HMI tags "Tool_Editor"
   "DB_MouldEditor_HMI_uData_sSelected_iCalculation" : Int = PLC DB_MouldEditor_HMI.uData.sSelected.iCalculation AT %DB10.DBW92, 1 s
   "DB_MouldEditor_HMI_uData_arShotSet{1}_CPMoveAfterShot" : Bool = PLC DB_MouldEditor_HMI.uData.arShotSet[1].CPMoveAfterShot AT %DB10.DBX236.1, 1 s
   "DB_MouldEditor_HMI_uData_arShotSet{2}_CPMoveAfterShot" : Bool = PLC DB_MouldEditor_HMI.uData.arShotSet[2].CPMoveAfterShot AT %DB10.DBX308.1, 1 s
   "DB_MouldEditor_HMI_uData_arShotSet{3}_CPMoveAfterShot" : Bool = PLC DB_MouldEditor_HMI.uData.arShotSet[3].CPMoveAfterShot AT %DB10.DBX380.1, 1 s
   "DB_MouldEditor_HMI_uData_arShotSet{4}_CPMoveAfterShot" : Bool = PLC DB_MouldEditor_HMI.uData.arShotSet[4].CPMoveAfterShot AT %DB10.DBX452.1, 1 s
   "DB_MouldEditor_HMI_uData_arShotSet{5}_CPMoveAfterShot" : Bool = PLC DB_MouldEditor_HMI.uData.arShotSet[5].CPMoveAfterShot AT %DB10.DBX524.1, 1 s
   "DB_MouldEditor_HMI_uData_arShotSet{6}_CPMoveAfterShot" : Bool = PLC DB_MouldEditor_HMI.uData.arShotSet[6].CPMoveAfterShot AT %DB10.DBX596.1, 1 s
   "DB_MouldEditor_HMI_uData_arShotSet{7}_CPMoveAfterShot" : Bool = PLC DB_MouldEditor_HMI.uData.arShotSet[7].CPMoveAfterShot AT %DB10.DBX668.1, 1 s
   "DB_MouldEditor_HMI_uData_arShotSet{8}_CPMoveAfterShot" : Bool = PLC DB_MouldEditor_HMI.uData.arShotSet[8].CPMoveAfterShot AT %DB10.DBX740.1, 1 s
   "DB_MouldEditor_HMI_uData_uTools_EnableTool" : Bool = PLC DB_MouldEditor_HMI.uData.uTools.EnableTool AT %DB10.DBX771.0, 1 s
   "DB_MouldEditor_HMI_uData_sSelected_sPS_arFlow{1}" : Real = PLC DB_MouldEditor_HMI.uData.sSelected.sPS.arFlow[1] AT %DB10.DBD8, 1 s
   "DB_MouldEditor_HMI_uData_sSelected_sPS_arFlow{2}" : Real = PLC DB_MouldEditor_HMI.uData.sSelected.sPS.arFlow[2] AT %DB10.DBD12, 1 s
   "DB_MouldEditor_HMI_uData_sSelected_sPS_arFlow{3}" : Real = PLC DB_MouldEditor_HMI.uData.sSelected.sPS.arFlow[3] AT %DB10.DBD16, 1 s
   "DB_MouldEditor_HMI_uData_sSelected_sPS_arFlow{4}" : Real = PLC DB_MouldEditor_HMI.uData.sSelected.sPS.arFlow[4] AT %DB10.DBD20, 1 s
   "DB_MouldEditor_HMI_uData_sSelected_sPS_arFlow{5}" : Real = PLC DB_MouldEditor_HMI.uData.sSelected.sPS.arFlow[5] AT %DB10.DBD24, 1 s
   "DB_MouldEditor_HMI_uData_sSelected_sPS_arFlow{6}" : Real = PLC DB_MouldEditor_HMI.uData.sSelected.sPS.arFlow[6] AT %DB10.DBD28, 1 s
   "DB_MouldEditor_HMI_uData_arShotSet{1}_MHNo" : Int = PLC DB_MouldEditor_HMI.uData.arShotSet[1].MHNo AT %DB10.DBW166, 1 s
   "DB_MouldEditor_HMI_uData_arShotSet{2}_MHNo" : Int = PLC DB_MouldEditor_HMI.uData.arShotSet[2].MHNo AT %DB10.DBW238, 1 s
   "DB_MouldEditor_HMI_uData_arShotSet{3}_MHNo" : Int = PLC DB_MouldEditor_HMI.uData.arShotSet[3].MHNo AT %DB10.DBW310, 1 s
   "DB_MouldEditor_HMI_uData_arShotSet{4}_MHNo" : Int = PLC DB_MouldEditor_HMI.uData.arShotSet[4].MHNo AT %DB10.DBW382, 1 s
   "DB_MouldEditor_HMI_uData_arShotSet{5}_MHNo" : Int = PLC DB_MouldEditor_HMI.uData.arShotSet[5].MHNo AT %DB10.DBW454, 1 s
   "DB_MouldEditor_HMI_uData_arShotSet{6}_MHNo" : Int = PLC DB_MouldEditor_HMI.uData.arShotSet[6].MHNo AT %DB10.DBW526, 1 s
   "DB_MouldEditor_HMI_uData_arShotSet{7}_MHNo" : Int = PLC DB_MouldEditor_HMI.uData.arShotSet[7].MHNo AT %DB10.DBW598, 1 s
   "DB_MouldEditor_HMI_uData_arShotSet{8}_MHNo" : Int = PLC DB_MouldEditor_HMI.uData.arShotSet[8].MHNo AT %DB10.DBW670, 1 s
   "DB_MouldEditor_HMI_uData_arShotSet{1}_PartCounter" : Int = PLC DB_MouldEditor_HMI.uData.arShotSet[1].PartCounter AT %DB10.DBW184, 1 s
   "DB_MouldEditor_HMI_uData_arShotSet{2}_PartCounter" : Int = PLC DB_MouldEditor_HMI.uData.arShotSet[2].PartCounter AT %DB10.DBW256, 1 s
   "DB_MouldEditor_HMI_uData_arShotSet{3}_PartCounter" : Int = PLC DB_MouldEditor_HMI.uData.arShotSet[3].PartCounter AT %DB10.DBW328, 1 s
   "DB_MouldEditor_HMI_uData_arShotSet{4}_PartCounter" : Int = PLC DB_MouldEditor_HMI.uData.arShotSet[4].PartCounter AT %DB10.DBW400, 1 s
   "DB_MouldEditor_HMI_uData_arShotSet{5}_PartCounter" : Int = PLC DB_MouldEditor_HMI.uData.arShotSet[5].PartCounter AT %DB10.DBW472, 1 s
   "DB_MouldEditor_HMI_uData_arShotSet{6}_PartCounter" : Int = PLC DB_MouldEditor_HMI.uData.arShotSet[6].PartCounter AT %DB10.DBW544, 1 s
   "DB_MouldEditor_HMI_uData_arShotSet{7}_PartCounter" : Int = PLC DB_MouldEditor_HMI.uData.arShotSet[7].PartCounter AT %DB10.DBW616, 1 s
   "DB_MouldEditor_HMI_uData_arShotSet{8}_PartCounter" : Int = PLC DB_MouldEditor_HMI.uData.arShotSet[8].PartCounter AT %DB10.DBW688, 1 s
   "DB_MouldEditor_HMI_uData_arShotSet{1}_PartWeight" : Real = PLC DB_MouldEditor_HMI.uData.arShotSet[1].PartWeight AT %DB10.DBD172, 1 s
   "DB_MouldEditor_HMI_uData_arShotSet{2}_PartWeight" : Real = PLC DB_MouldEditor_HMI.uData.arShotSet[2].PartWeight AT %DB10.DBD244, 1 s
   "DB_MouldEditor_HMI_uData_arShotSet{3}_PartWeight" : Real = PLC DB_MouldEditor_HMI.uData.arShotSet[3].PartWeight AT %DB10.DBD316, 1 s
   "DB_MouldEditor_HMI_uData_arShotSet{4}_PartWeight" : Real = PLC DB_MouldEditor_HMI.uData.arShotSet[4].PartWeight AT %DB10.DBD388, 1 s
   "DB_MouldEditor_HMI_uData_arShotSet{5}_PartWeight" : Real = PLC DB_MouldEditor_HMI.uData.arShotSet[5].PartWeight AT %DB10.DBD460, 1 s
   "DB_MouldEditor_HMI_uData_arShotSet{6}_PartWeight" : Real = PLC DB_MouldEditor_HMI.uData.arShotSet[6].PartWeight AT %DB10.DBD532, 1 s
   "DB_MouldEditor_HMI_uData_arShotSet{7}_PartWeight" : Real = PLC DB_MouldEditor_HMI.uData.arShotSet[7].PartWeight AT %DB10.DBD604, 1 s
   "DB_MouldEditor_HMI_uData_arShotSet{8}_PartWeight" : Real = PLC DB_MouldEditor_HMI.uData.arShotSet[8].PartWeight AT %DB10.DBD676, 1 s
   "DB_MouldEditor_HMI_uData_sSelected_sPS_arPressure{1}" : Real = PLC DB_MouldEditor_HMI.uData.sSelected.sPS.arPressure[1] AT %DB10.DBD64, 1 s
   "DB_MouldEditor_HMI_uData_sSelected_sPS_arPressure{2}" : Real = PLC DB_MouldEditor_HMI.uData.sSelected.sPS.arPressure[2] AT %DB10.DBD68, 1 s
   "DB_MouldEditor_HMI_uData_sSelected_sPS_arPressure{3}" : Real = PLC DB_MouldEditor_HMI.uData.sSelected.sPS.arPressure[3] AT %DB10.DBD72, 1 s
   "DB_MouldEditor_HMI_uData_sSelected_sPS_arPressure{4}" : Real = PLC DB_MouldEditor_HMI.uData.sSelected.sPS.arPressure[4] AT %DB10.DBD76, 1 s
   "DB_MouldEditor_HMI_uData_sSelected_sPS_arPressure{5}" : Real = PLC DB_MouldEditor_HMI.uData.sSelected.sPS.arPressure[5] AT %DB10.DBD80, 1 s
   "DB_MouldEditor_HMI_uData_sSelected_sPS_arPressure{6}" : Real = PLC DB_MouldEditor_HMI.uData.sSelected.sPS.arPressure[6] AT %DB10.DBD84, 1 s
   "DB_MouldEditor_HMI_uData_arShotSet{1}_PartShotDisable" : Bool = PLC DB_MouldEditor_HMI.uData.arShotSet[1].PartShotDisable AT %DB10.DBX236.0, 1 s
   "DB_MouldEditor_HMI_uData_arShotSet{2}_PartShotDisable" : Bool = PLC DB_MouldEditor_HMI.uData.arShotSet[2].PartShotDisable AT %DB10.DBX308.0, 1 s
   "DB_MouldEditor_HMI_uData_arShotSet{3}_PartShotDisable" : Bool = PLC DB_MouldEditor_HMI.uData.arShotSet[3].PartShotDisable AT %DB10.DBX380.0, 1 s
   "DB_MouldEditor_HMI_uData_arShotSet{4}_PartShotDisable" : Bool = PLC DB_MouldEditor_HMI.uData.arShotSet[4].PartShotDisable AT %DB10.DBX452.0, 1 s
   "DB_MouldEditor_HMI_uData_arShotSet{5}_PartShotDisable" : Bool = PLC DB_MouldEditor_HMI.uData.arShotSet[5].PartShotDisable AT %DB10.DBX524.0, 1 s
   "DB_MouldEditor_HMI_uData_arShotSet{6}_PartShotDisable" : Bool = PLC DB_MouldEditor_HMI.uData.arShotSet[6].PartShotDisable AT %DB10.DBX596.0, 1 s
   "DB_MouldEditor_HMI_uData_arShotSet{7}_PartShotDisable" : Bool = PLC DB_MouldEditor_HMI.uData.arShotSet[7].PartShotDisable AT %DB10.DBX668.0, 1 s
   "DB_MouldEditor_HMI_uData_arShotSet{8}_PartShotDisable" : Bool = PLC DB_MouldEditor_HMI.uData.arShotSet[8].PartShotDisable AT %DB10.DBX740.0, 1 s
   "DB_MouldEditor_HMI_uData_sSelected_sPS_iPS" : Int = PLC DB_MouldEditor_HMI.uData.sSelected.sPS.iPS AT %DB10.DBW2, 1 s
   "DB_MouldEditor_HMI_uData_sSelected_sPS_arRatio{1}" : Real = PLC DB_MouldEditor_HMI.uData.sSelected.sPS.arRatio[1] AT %DB10.DBD36, 1 s
   "DB_MouldEditor_HMI_uData_sSelected_sPS_arRatio{2}" : Real = PLC DB_MouldEditor_HMI.uData.sSelected.sPS.arRatio[2] AT %DB10.DBD40, 1 s
   "DB_MouldEditor_HMI_uData_sSelected_sPS_arRatio{3}" : Real = PLC DB_MouldEditor_HMI.uData.sSelected.sPS.arRatio[3] AT %DB10.DBD44, 1 s
   "DB_MouldEditor_HMI_uData_sSelected_sPS_arRatio{4}" : Real = PLC DB_MouldEditor_HMI.uData.sSelected.sPS.arRatio[4] AT %DB10.DBD48, 1 s
   "DB_MouldEditor_HMI_uData_sSelected_sPS_arRatio{5}" : Real = PLC DB_MouldEditor_HMI.uData.sSelected.sPS.arRatio[5] AT %DB10.DBD52, 1 s
   "DB_MouldEditor_HMI_uData_sSelected_sPS_arRatio{6}" : Real = PLC DB_MouldEditor_HMI.uData.sSelected.sPS.arRatio[6] AT %DB10.DBD56, 1 s
   "DB_MouldEditor_HMI_uData_arShotSet{1}_PurgeMHAfterShot" : Bool = PLC DB_MouldEditor_HMI.uData.arShotSet[1].PurgeMHAfterShot AT %DB10.DBX236.2, 1 s
   "DB_MouldEditor_HMI_uData_arShotSet{2}_PurgeMHAfterShot" : Bool = PLC DB_MouldEditor_HMI.uData.arShotSet[2].PurgeMHAfterShot AT %DB10.DBX308.2, 1 s
   "DB_MouldEditor_HMI_uData_arShotSet{3}_PurgeMHAfterShot" : Bool = PLC DB_MouldEditor_HMI.uData.arShotSet[3].PurgeMHAfterShot AT %DB10.DBX380.2, 1 s
   "DB_MouldEditor_HMI_uData_arShotSet{4}_PurgeMHAfterShot" : Bool = PLC DB_MouldEditor_HMI.uData.arShotSet[4].PurgeMHAfterShot AT %DB10.DBX452.2, 1 s
   "DB_MouldEditor_HMI_uData_arShotSet{5}_PurgeMHAfterShot" : Bool = PLC DB_MouldEditor_HMI.uData.arShotSet[5].PurgeMHAfterShot AT %DB10.DBX524.2, 1 s
   "DB_MouldEditor_HMI_uData_arShotSet{6}_PurgeMHAfterShot" : Bool = PLC DB_MouldEditor_HMI.uData.arShotSet[6].PurgeMHAfterShot AT %DB10.DBX596.2, 1 s
   "DB_MouldEditor_HMI_uData_arShotSet{7}_PurgeMHAfterShot" : Bool = PLC DB_MouldEditor_HMI.uData.arShotSet[7].PurgeMHAfterShot AT %DB10.DBX668.2, 1 s
   "DB_MouldEditor_HMI_uData_arShotSet{8}_PurgeMHAfterShot" : Bool = PLC DB_MouldEditor_HMI.uData.arShotSet[8].PurgeMHAfterShot AT %DB10.DBX740.2, 1 s
   "DB_MouldEditor_HMI_uData_arShotSet{1}_FoamingTime" : Real = PLC DB_MouldEditor_HMI.uData.arShotSet[1].FoamingTime AT %DB10.DBD168, 1 s
   "DB_MouldEditor_HMI_uData_arShotSet{2}_FoamingTime" : Real = PLC DB_MouldEditor_HMI.uData.arShotSet[2].FoamingTime AT %DB10.DBD240, 1 s
   "DB_MouldEditor_HMI_uData_arShotSet{3}_FoamingTime" : Real = PLC DB_MouldEditor_HMI.uData.arShotSet[3].FoamingTime AT %DB10.DBD312, 1 s
   "DB_MouldEditor_HMI_uData_arShotSet{4}_FoamingTime" : Real = PLC DB_MouldEditor_HMI.uData.arShotSet[4].FoamingTime AT %DB10.DBD384, 1 s
   "DB_MouldEditor_HMI_uData_arShotSet{5}_FoamingTime" : Real = PLC DB_MouldEditor_HMI.uData.arShotSet[5].FoamingTime AT %DB10.DBD456, 1 s
   "DB_MouldEditor_HMI_uData_arShotSet{6}_FoamingTime" : Real = PLC DB_MouldEditor_HMI.uData.arShotSet[6].FoamingTime AT %DB10.DBD528, 1 s
   "DB_MouldEditor_HMI_uData_arShotSet{7}_FoamingTime" : Real = PLC DB_MouldEditor_HMI.uData.arShotSet[7].FoamingTime AT %DB10.DBD600, 1 s
   "DB_MouldEditor_HMI_uData_arShotSet{8}_FoamingTime" : Real = PLC DB_MouldEditor_HMI.uData.arShotSet[8].FoamingTime AT %DB10.DBD672, 1 s
   "DB_MouldEditor_HMI_uData_uTools_tool_name" : String[20] = PLC DB_MouldEditor_HMI.uData.uTools.tool_name AT %DB10.DBX742.0, 1 s
   "DB_MouldEditor_HMI_uData_sCalculatedValues_arTotalFlow{1}" : Real = PLC DB_MouldEditor_HMI.uData.sCalculatedValues.arTotalFlow[1] AT %DB10.DBD780, 1 s
   "DB_MouldEditor_HMI_uData_sCalculatedValues_arTotalFlow{2}" : Real = PLC DB_MouldEditor_HMI.uData.sCalculatedValues.arTotalFlow[2] AT %DB10.DBD784, 1 s
   "DB_MouldEditor_HMI_uData_sCalculatedValues_arTotalFlow{3}" : Real = PLC DB_MouldEditor_HMI.uData.sCalculatedValues.arTotalFlow[3] AT %DB10.DBD788, 1 s
   "DB_MouldEditor_HMI_uData_sCalculatedValues_arTotalFlow{4}" : Real = PLC DB_MouldEditor_HMI.uData.sCalculatedValues.arTotalFlow[4] AT %DB10.DBD792, 1 s
   "DB_MouldEditor_HMI_uData_sCalculatedValues_arTotalFlow{5}" : Real = PLC DB_MouldEditor_HMI.uData.sCalculatedValues.arTotalFlow[5] AT %DB10.DBD796, 1 s
   "DB_MouldEditor_HMI_uData_sCalculatedValues_arTotalFlow{6}" : Real = PLC DB_MouldEditor_HMI.uData.sCalculatedValues.arTotalFlow[6] AT %DB10.DBD800, 1 s
   "DB_MouldEditor_HMI_uData_sCalculatedValues_arTotalFlow{7}" : Real = PLC DB_MouldEditor_HMI.uData.sCalculatedValues.arTotalFlow[7] AT %DB10.DBD804, 1 s
   "DB_MouldEditor_HMI_uData_sCalculatedValues_arTotalFlow{8}" : Real = PLC DB_MouldEditor_HMI.uData.sCalculatedValues.arTotalFlow[8] AT %DB10.DBD808, 1 s
   "DB_MouldEditor_HMI_uData_uTools_PartShot_Amount" : Byte = PLC DB_MouldEditor_HMI.uData.uTools.PartShot_Amount AT %DB10.DBB768, 1 s
   "DB_MouldEditor_HMI_uData_sStatusBits_xValueChanged" : Bool = PLC DB_MouldEditor_HMI.uData.sStatusBits.xValueChanged AT %DB10.DBX812.0, 1 s
   "DB_MouldEditor_HMI_uData_sStatusBits_xSafeChanges" : Bool = PLC DB_MouldEditor_HMI.uData.sStatusBits.xSafeChanges AT %DB10.DBX812.1, 1 s
   "DB_MouldEditor_HMI_uData_sStatusBits_xDiscardChanges" : Bool = PLC DB_MouldEditor_HMI.uData.sStatusBits.xDiscardChanges AT %DB10.DBX812.2, 1 s
   "DB_MouldEditor_HMI_uData_sStatusBits_xDeleteProgram" : Bool = PLC DB_MouldEditor_HMI.uData.sStatusBits.xDeleteProgram AT %DB10.DBX812.3, 1 s
   "DB_MouldEditor_HMI_uData_sStatusBits_xFaultDeleteProgram" : Bool = PLC DB_MouldEditor_HMI.uData.sStatusBits.xFaultDeleteProgram AT %DB10.DBX812.4, 1 s
      on ChangeValue: "PopUp_ToolEditor"()
   "DB_MouldEditor_HMI_uData_sStatusBits_xProgLoadName" : Bool = PLC DB_MouldEditor_HMI.uData.sStatusBits.xProgLoadName AT %DB10.DBX812.5, 1 s
   "DB_MouldEditor_HMI_uData_sStatusBits_xProgLoadNameAckn" : Bool = PLC DB_MouldEditor_HMI.uData.sStatusBits.xProgLoadNameAckn AT %DB10.DBX812.6, 1 s
   "DB_MouldEditor_HMI_uData_sStatusBits_xFaultValuesnotvalid" : Bool = PLC DB_MouldEditor_HMI.uData.sStatusBits.xFaultValuesnotvalid AT %DB10.DBX812.7, 1 s
      on ChangeValue: "Show_Not_Valid"()
   "DB_MouldEditor_HMI_uData_sStatusBits_xPartShotAmount_increase" : Bool = PLC DB_MouldEditor_HMI.uData.sStatusBits.xPartShotAmount_increase AT %DB10.DBX813.0, 1 s
   "DB_MouldEditor_HMI_uData_sStatusBits_xPartShotAmount_decrease" : Bool = PLC DB_MouldEditor_HMI.uData.sStatusBits.xPartShotAmount_decrease AT %DB10.DBX813.1, 1 s
   "Activate_Deactivate" : Bool AT %DB1.DBB0
   "Coloum_Activate" : Int, internal
   "InterfaceVisu_ReadWriteDeviceNo" : Int = PLC InterfaceVisu.ReadWriteDeviceNo AT %DB1.DBW100, 1 s
   "DB_MouldEditor_HMI_uData_sSelected_iTool" : Int = PLC DB_MouldEditor_HMI.uData.sSelected.iTool AT %DB10.DBW0, 1 s
   "DB_MouldEditor_HMI_uData_sSelected_sPS_RefComponent" : Int = PLC DB_MouldEditor_HMI.uData.sSelected.sPS.RefComponent AT %DB10.DBW88, 1 s
   "InterfaceVisu_SetHDValue" : Bool = PLC InterfaceVisu.SetHDValue AT %DB1.DBX104.4, 1 s
   "DB_MouldEditor_HMI_uData_uTools_Rob_Prog" : Int = PLC DB_MouldEditor_HMI.uData.uTools.Rob_Prog AT %DB10.DBW764, 1 s
   "DB_MouldEditor_HMI_uData_uTools_Rob_Prog2" : Int = PLC DB_MouldEditor_HMI.uData.uTools.Rob_Prog2 AT %DB10.DBW766, 1 s
   "DB_MouldEditor_HMI_uData_uTools_Spare" : Byte = PLC DB_MouldEditor_HMI.uData.uTools.Spare AT %DB10.DBB770, 1 s
   "DB_MouldEditor_HMI_uData_uTools_Spare5_2" : Bool = PLC DB_MouldEditor_HMI.uData.uTools.Spare5_2 AT %DB10.DBX771.1, 1 s
   "DB_MouldEditor_HMI_uData_uTools_Spare5_3" : Bool = PLC PN_Mixinghead.Mixinghead[0].DüseBypass[4].Visualisierung.OutputForNozzle AT %DB10.DBX771.2, 1 s
   "DB_MouldEditor_HMI_uData_uTools_Spare5_4" : Bool = PLC DB_MouldEditor_HMI.uData.uTools.Spare5_4 AT %DB10.DBX771.3, 1 s
   "DB_MouldEditor_HMI_uData_uTools_Spare5_5" : Bool = PLC DB_MouldEditor_HMI.uData.uTools.Spare5_5 AT %DB10.DBX771.4, 1 s
   "DB_MouldEditor_HMI_uData_uTools_Spare5_6" : Bool = PLC DB_MouldEditor_HMI.uData.uTools.Spare5_6 AT %DB10.DBX771.5, 1 s
   "DB_MouldEditor_HMI_uData_uTools_EnablePurgeMH" : Bool = PLC DB_MouldEditor_HMI.uData.uTools.EnablePurgeMH AT %DB10.DBX771.6, 1 s
   "DB_MouldEditor_HMI_uData_uTools_NitrogenVol" : Int = PLC DB_MouldEditor_HMI.uData.uTools.NitrogenVol AT %DB10.DBW772, 1 s
   "DB_MouldEditor_HMI_uData_uTools_Spare_12" : Word = PLC DB_MouldEditor_HMI.uData.uTools.Spare_12 AT %DB10.DBW774, 1 s
   "DB_MouldEditor_HMI_uData_uTools_RefComponent" : Byte = PLC DB_MouldEditor_HMI.uData.uTools.RefComponent AT %DB10.DBB769, 1 s
   "DB_MouldEditor_HMI_uData_sColumn_iShotTime" : Int = PLC DB612_Tank_State.Tank[2].Max_Level AT %DB10.DBW814, 1 s
   "DB_MouldEditor_HMI_uData_sColumn_iTotalFlow" : Int = PLC DB_MouldEditor_HMI.uData.sColumn.iTotalFlow AT %DB10.DBW816, 1 s
   "DB_MouldEditor_HMI_uData_sColumn_iTotalWeight" : Int = PLC DB_MouldEditor_HMI.uData.sColumn.iTotalWeight AT %DB10.DBW818, 1 s
   "DB_MouldEditor_HMI_uData_sRow_arChangePartialShot{0}" : Bool = PLC DB_MouldEditor_HMI.uData.sRow.arChangePartialShot[0] AT %DB10.DBX820.0, 1 s
   "DB_MouldEditor_HMI_uData_sRow_arChangePartialShot{1}" : Bool = PLC DB_MouldEditor_HMI.uData.sRow.arChangePartialShot[1] AT %DB10.DBX820.1, 1 s
   "DB_MouldEditor_HMI_uData_sRow_arChangePartialShot{2}" : Bool = PLC DB_MouldEditor_HMI.uData.sRow.arChangePartialShot[2] AT %DB10.DBX820.2, 1 s
   "DB_MouldEditor_HMI_uData_sRow_arChangePartialShot{3}" : Bool = PLC DB_MouldEditor_HMI.uData.sRow.arChangePartialShot[3] AT %DB10.DBX820.3, 1 s
   "DB_MouldEditor_HMI_uData_sRow_arChangePartialShot{4}" : Bool = PLC DB_MouldEditor_HMI.uData.sRow.arChangePartialShot[4] AT %DB10.DBX820.4, 1 s
   "DB_MouldEditor_HMI_uData_sRow_arChangePartialShot{5}" : Bool = PLC DB_MouldEditor_HMI.uData.sRow.arChangePartialShot[5] AT %DB10.DBX820.5, 1 s
   "DB_MouldEditor_HMI_uData_sRow_arChangePartialShot{6}" : Bool = PLC DB_MouldEditor_HMI.uData.sRow.arChangePartialShot[6] AT %DB10.DBX820.6, 1 s
   "DB_MouldEditor_HMI_uData_sRow_arChangePartialShot{7}" : Bool = PLC DB_MouldEditor_HMI.uData.sRow.arChangePartialShot[7] AT %DB10.DBX820.7, 1 s
   "DB_MouldEditor_HMI_uData_sRow_arChangePartialShot{8}" : Bool = PLC DB_MouldEditor_HMI.uData.sRow.arChangePartialShot[8] AT %DB10.DBX821.0, 1 s
   "DB_MouldEditor_HMI_uData_sCalculatedValues_arTotalFlow{0}" : Real = PLC DB_MouldEditor_HMI.uData.sCalculatedValues.arTotalFlow[0] AT %DB10.DBD776, 1 s
   "DB_MouldEditor_HMI_uData_arShotSet{0}_MHNo" : Int = PLC DB_MouldEditor_HMI.uData.arShotSet[0].MHNo AT %DB10.DBW94, 1 s
   "DB_MouldEditor_HMI_uData_arShotSet{0}_FoamingTime" : Real = PLC DB_MouldEditor_HMI.uData.arShotSet[0].FoamingTime AT %DB10.DBD96, 1 s
   "DB_MouldEditor_HMI_uData_arShotSet{0}_PartWeight" : Real = PLC DB_MouldEditor_HMI.uData.arShotSet[0].PartWeight AT %DB10.DBD100, 1 s
   "DB_MouldEditor_HMI_uData_arShotSet{0}_CP_ThrottleGap" : Real = PLC DB_MouldEditor_HMI.uData.arShotSet[0].CP_ThrottleGap AT %DB10.DBD104, 1 s
   "DB_MouldEditor_HMI_uData_arShotSet{0}_SwitchOff_Pressure" : Real = PLC DB_MouldEditor_HMI.uData.arShotSet[0].SwitchOff_Pressure AT %DB10.DBD108, 1 s
   "DB_MouldEditor_HMI_uData_arShotSet{0}_PartCounter" : Int = PLC DB_MouldEditor_HMI.uData.arShotSet[0].PartCounter AT %DB10.DBW112, 1 s
   "DB_MouldEditor_HMI_uData_arShotSet{0}_RefComponent" : Int = PLC DB_MouldEditor_HMI.uData.arShotSet[0].RefComponent AT %DB10.DBW162, 1 s
   "DB_MouldEditor_HMI_uData_arShotSet{0}_PartShotDisable" : Bool = PLC DB_MouldEditor_HMI.uData.arShotSet[0].PartShotDisable AT %DB10.DBX164.0, 1 s
   "DB_MouldEditor_HMI_uData_arShotSet{0}_CPMoveAfterShot" : Bool = PLC DB_MouldEditor_HMI.uData.arShotSet[0].CPMoveAfterShot AT %DB10.DBX164.1, 1 s
   "DB_MouldEditor_HMI_uData_arShotSet{0}_PurgeMHAfterShot" : Bool = PLC DB_MouldEditor_HMI.uData.arShotSet[0].PurgeMHAfterShot AT %DB10.DBX164.2, 1 s
   "DB_MouldEditor_HMI_uData_arShotSet{0}_2PoinMovement_Comp01" : Bool = PLC DB_MouldEditor_HMI.uData.arShotSet[0].2PoinMovement_Comp01 AT %DB10.DBX164.3, 1 s
   "DB_MouldEditor_HMI_uData_arShotSet{0}_2PoinMovement_Comp02" : Bool = PLC DB_MouldEditor_HMI.uData.arShotSet[0].2PoinMovement_Comp02 AT %DB10.DBX164.4, 1 s
   "DB_MouldEditor_HMI_uData_arShotSet{0}_2PoinMovement_Comp03" : Bool = PLC DB_MouldEditor_HMI.uData.arShotSet[0].2PoinMovement_Comp03 AT %DB10.DBX164.5, 1 s
   "DB_MouldEditor_HMI_uData_arShotSet{0}_2PoinMovement_Comp04" : Bool = PLC DB_MouldEditor_HMI.uData.arShotSet[0].2PoinMovement_Comp04 AT %DB10.DBX164.6, 1 s
   "DB_MouldEditor_HMI_uData_arShotSet{0}_2PoinMovement_Comp05" : Bool = PLC DB_MouldEditor_HMI.uData.arShotSet[0].2PoinMovement_Comp05 AT %DB10.DBX164.7, 1 s
   "DB_MouldEditor_HMI_uData_arShotSet{0}_2PoinMovement_Comp06" : Bool = PLC DB_MouldEditor_HMI.uData.arShotSet[0].2PoinMovement_Comp06 AT %DB10.DBX165.0, 1 s
   "DB_MouldEditor_HMI_uData_arShotSet{0}_Spare_1" : Bool = PLC DB_MouldEditor_HMI.uData.arShotSet[0].Spare_1 AT %DB10.DBX165.1, 1 s
   "DB_MouldEditor_HMI_uData_arShotSet{0}_Spare_2" : Bool = PLC DB_MouldEditor_HMI.uData.arShotSet[0].Spare_2 AT %DB10.DBX165.2, 1 s
   "DB_MouldEditor_HMI_uData_arShotSet{0}_Spare_3" : Bool = PLC DB_MouldEditor_HMI.uData.arShotSet[0].Spare_3 AT %DB10.DBX165.3, 1 s
   "DB_MouldEditor_HMI_uData_arShotSet{0}_Spare_4" : Bool = PLC DB_MouldEditor_HMI.uData.arShotSet[0].Spare_4 AT %DB10.DBX165.4, 1 s
   "DB_MouldEditor_HMI_uData_arShotSet{0}_Spare_5" : Bool = PLC DB_MouldEditor_HMI.uData.arShotSet[0].Spare_5 AT %DB10.DBX165.5, 1 s
   "DB_MouldEditor_HMI_uData_arShotSet{0}_Spare_6" : Bool = PLC DB_MouldEditor_HMI.uData.arShotSet[0].Spare_6 AT %DB10.DBX165.6, 1 s
   "DB_MouldEditor_HMI_uData_arShotSet{0}_Spare_7" : Bool = PLC DB_MouldEditor_HMI.uData.arShotSet[0].Spare_7 AT %DB10.DBX165.7, 1 s
   "DB_MouldEditor_HMI_uData_arShotSet{1}_CP_ThrottleGap" : Real = PLC DB_MouldEditor_HMI.uData.arShotSet[1].CP_ThrottleGap AT %DB10.DBD176, 1 s
   "DB_MouldEditor_HMI_uData_arShotSet{1}_SwitchOff_Pressure" : Real = PLC DB_MouldEditor_HMI.uData.arShotSet[1].SwitchOff_Pressure AT %DB10.DBD180, 1 s
   "DB_MouldEditor_HMI_uData_arShotSet{1}_RefComponent" : Int = PLC DB_MouldEditor_HMI.uData.arShotSet[1].RefComponent AT %DB10.DBW234, 1 s
   "DB_MouldEditor_HMI_uData_arShotSet{1}_2PoinMovement_Comp01" : Bool = PLC DB_MouldEditor_HMI.uData.arShotSet[1].2PoinMovement_Comp01 AT %DB10.DBX236.3, 1 s
   "DB_MouldEditor_HMI_uData_arShotSet{1}_2PoinMovement_Comp02" : Bool = PLC DB_MouldEditor_HMI.uData.arShotSet[1].2PoinMovement_Comp02 AT %DB10.DBX236.4, 1 s
   "DB_MouldEditor_HMI_uData_arShotSet{1}_2PoinMovement_Comp03" : Bool = PLC DB_MouldEditor_HMI.uData.arShotSet[1].2PoinMovement_Comp03 AT %DB10.DBX236.5, 1 s
   "DB_MouldEditor_HMI_uData_arShotSet{1}_2PoinMovement_Comp04" : Bool = PLC DB_MouldEditor_HMI.uData.arShotSet[1].2PoinMovement_Comp04 AT %DB10.DBX236.6, 1 s
   "DB_MouldEditor_HMI_uData_arShotSet{1}_2PoinMovement_Comp05" : Bool = PLC DB_MouldEditor_HMI.uData.arShotSet[1].2PoinMovement_Comp05 AT %DB10.DBX236.7, 1 s
   "DB_MouldEditor_HMI_uData_arShotSet{1}_2PoinMovement_Comp06" : Bool = PLC DB_MouldEditor_HMI.uData.arShotSet[1].2PoinMovement_Comp06 AT %DB10.DBX237.0, 1 s
   "DB_MouldEditor_HMI_uData_arShotSet{1}_Spare_1" : Bool = PLC DB_MouldEditor_HMI.uData.arShotSet[1].Spare_1 AT %DB10.DBX237.1, 1 s
   "DB_MouldEditor_HMI_uData_arShotSet{1}_Spare_2" : Bool = PLC DB_MouldEditor_HMI.uData.arShotSet[1].Spare_2 AT %DB10.DBX237.2, 1 s
   "DB_MouldEditor_HMI_uData_arShotSet{1}_Spare_3" : Bool = PLC DB_MouldEditor_HMI.uData.arShotSet[1].Spare_3 AT %DB10.DBX237.3, 1 s
   "DB_MouldEditor_HMI_uData_arShotSet{1}_Spare_4" : Bool = PLC DB_MouldEditor_HMI.uData.arShotSet[1].Spare_4 AT %DB10.DBX237.4, 1 s
   "DB_MouldEditor_HMI_uData_arShotSet{1}_Spare_5" : Bool = PLC DB_MouldEditor_HMI.uData.arShotSet[1].Spare_5 AT %DB10.DBX237.5, 1 s
   "DB_MouldEditor_HMI_uData_arShotSet{1}_Spare_6" : Bool = PLC DB_MouldEditor_HMI.uData.arShotSet[1].Spare_6 AT %DB10.DBX237.6, 1 s
   "DB_MouldEditor_HMI_uData_arShotSet{1}_Spare_7" : Bool = PLC DB_MouldEditor_HMI.uData.arShotSet[1].Spare_7 AT %DB10.DBX237.7, 1 s
   "DB_MouldEditor_HMI_uData_arShotSet{2}_CP_ThrottleGap" : Real = PLC DB_MouldEditor_HMI.uData.arShotSet[2].CP_ThrottleGap AT %DB10.DBD248, 1 s
   "DB_MouldEditor_HMI_uData_arShotSet{2}_SwitchOff_Pressure" : Real = PLC DB_MouldEditor_HMI.uData.arShotSet[2].SwitchOff_Pressure AT %DB10.DBD252, 1 s
   "DB_MouldEditor_HMI_uData_arShotSet{2}_RefComponent" : Int = PLC DB_MouldEditor_HMI.uData.arShotSet[2].RefComponent AT %DB10.DBW306, 1 s
   "DB_MouldEditor_HMI_uData_arShotSet{2}_2PoinMovement_Comp01" : Bool = PLC DB_MouldEditor_HMI.uData.arShotSet[2].2PoinMovement_Comp01 AT %DB10.DBX308.3, 1 s
   "DB_MouldEditor_HMI_uData_arShotSet{2}_2PoinMovement_Comp02" : Bool = PLC DB_MouldEditor_HMI.uData.arShotSet[2].2PoinMovement_Comp02 AT %DB10.DBX308.4, 1 s
   "DB_MouldEditor_HMI_uData_arShotSet{2}_2PoinMovement_Comp03" : Bool = PLC DB_MouldEditor_HMI.uData.arShotSet[2].2PoinMovement_Comp03 AT %DB10.DBX308.5, 1 s
   "DB_MouldEditor_HMI_uData_arShotSet{2}_2PoinMovement_Comp04" : Bool = PLC DB_MouldEditor_HMI.uData.arShotSet[2].2PoinMovement_Comp04 AT %DB10.DBX308.6, 1 s
   "DB_MouldEditor_HMI_uData_arShotSet{2}_2PoinMovement_Comp05" : Bool = PLC DB_MouldEditor_HMI.uData.arShotSet[2].2PoinMovement_Comp05 AT %DB10.DBX308.7, 1 s
   "DB_MouldEditor_HMI_uData_arShotSet{2}_2PoinMovement_Comp06" : Bool = PLC DB_MouldEditor_HMI.uData.arShotSet[2].2PoinMovement_Comp06 AT %DB10.DBX309.0, 1 s
   "DB_MouldEditor_HMI_uData_arShotSet{2}_Spare_1" : Bool = PLC DB_MouldEditor_HMI.uData.arShotSet[2].Spare_1 AT %DB10.DBX309.1, 1 s
   "DB_MouldEditor_HMI_uData_arShotSet{2}_Spare_2" : Bool = PLC DB_MouldEditor_HMI.uData.arShotSet[2].Spare_2 AT %DB10.DBX309.2, 1 s
   "DB_MouldEditor_HMI_uData_arShotSet{2}_Spare_3" : Bool = PLC DB_MouldEditor_HMI.uData.arShotSet[2].Spare_3 AT %DB10.DBX309.3, 1 s
   "DB_MouldEditor_HMI_uData_arShotSet{2}_Spare_4" : Bool = PLC DB_MouldEditor_HMI.uData.arShotSet[2].Spare_4 AT %DB10.DBX309.4, 1 s
   "DB_MouldEditor_HMI_uData_arShotSet{2}_Spare_5" : Bool = PLC DB_MouldEditor_HMI.uData.arShotSet[2].Spare_5 AT %DB10.DBX309.5, 1 s
   "DB_MouldEditor_HMI_uData_arShotSet{2}_Spare_6" : Bool = PLC DB_MouldEditor_HMI.uData.arShotSet[2].Spare_6 AT %DB10.DBX309.6, 1 s
   "DB_MouldEditor_HMI_uData_arShotSet{2}_Spare_7" : Bool = PLC DB_MouldEditor_HMI.uData.arShotSet[2].Spare_7 AT %DB10.DBX309.7, 1 s
   "DB_MouldEditor_HMI_uData_arShotSet{3}_CP_ThrottleGap" : Real = PLC DB602_PV_Tank.Tank[0].Level.PV_ActV.Value AT %DB10.DBD320, 1 s
   "DB_MouldEditor_HMI_uData_arShotSet{3}_SwitchOff_Pressure" : Real = PLC DB_MouldEditor_HMI.uData.arShotSet[3].SwitchOff_Pressure AT %DB10.DBD324, 1 s
   "DB_MouldEditor_HMI_uData_arShotSet{3}_RefComponent" : Int = PLC DB_MouldEditor_HMI.uData.arShotSet[3].RefComponent AT %DB10.DBW378, 1 s
   "DB_MouldEditor_HMI_uData_arShotSet{3}_2PoinMovement_Comp01" : Bool = PLC DB_MouldEditor_HMI.uData.arShotSet[3].2PoinMovement_Comp01 AT %DB10.DBX380.3, 1 s
   "DB_MouldEditor_HMI_uData_arShotSet{3}_2PoinMovement_Comp02" : Bool = PLC DB_MouldEditor_HMI.uData.arShotSet[3].2PoinMovement_Comp02 AT %DB10.DBX380.4, 1 s
   "DB_MouldEditor_HMI_uData_arShotSet{3}_2PoinMovement_Comp03" : Bool = PLC DB_MouldEditor_HMI.uData.arShotSet[3].2PoinMovement_Comp03 AT %DB10.DBX380.5, 1 s
   "DB_MouldEditor_HMI_uData_arShotSet{3}_2PoinMovement_Comp04" : Bool = PLC DB_MouldEditor_HMI.uData.arShotSet[3].2PoinMovement_Comp04 AT %DB10.DBX380.6, 1 s
   "DB_MouldEditor_HMI_uData_arShotSet{3}_2PoinMovement_Comp05" : Bool = PLC DB_MouldEditor_HMI.uData.arShotSet[3].2PoinMovement_Comp05 AT %DB10.DBX380.7, 1 s
   "DB_MouldEditor_HMI_uData_arShotSet{3}_2PoinMovement_Comp06" : Bool = PLC DB_MouldEditor_HMI.uData.arShotSet[3].2PoinMovement_Comp06 AT %DB10.DBX381.0, 1 s
   "DB_MouldEditor_HMI_uData_arShotSet{3}_Spare_1" : Bool = PLC DB_MouldEditor_HMI.uData.arShotSet[3].Spare_1 AT %DB10.DBX381.1, 1 s
   "DB_MouldEditor_HMI_uData_arShotSet{3}_Spare_2" : Bool = PLC DB_MouldEditor_HMI.uData.arShotSet[3].Spare_2 AT %DB10.DBX381.2, 1 s
   "DB_MouldEditor_HMI_uData_arShotSet{3}_Spare_3" : Bool = PLC DB_MouldEditor_HMI.uData.arShotSet[3].Spare_3 AT %DB10.DBX381.3, 1 s
   "DB_MouldEditor_HMI_uData_arShotSet{3}_Spare_4" : Bool = PLC DB_MouldEditor_HMI.uData.arShotSet[3].Spare_4 AT %DB10.DBX381.4, 1 s
   "DB_MouldEditor_HMI_uData_arShotSet{3}_Spare_5" : Bool = PLC DB_MouldEditor_HMI.uData.arShotSet[3].Spare_5 AT %DB10.DBX381.5, 1 s
   "DB_MouldEditor_HMI_uData_arShotSet{3}_Spare_6" : Bool = PLC DB_MouldEditor_HMI.uData.arShotSet[3].Spare_6 AT %DB10.DBX381.6, 1 s
   "DB_MouldEditor_HMI_uData_arShotSet{3}_Spare_7" : Bool = PLC DB_MouldEditor_HMI.uData.arShotSet[3].Spare_7 AT %DB10.DBX381.7, 1 s
   "DB_MouldEditor_HMI_uData_arShotSet{4}_CP_ThrottleGap" : Real = PLC DB_MouldEditor_HMI.uData.arShotSet[4].CP_ThrottleGap AT %DB10.DBD392, 1 s
   "DB_MouldEditor_HMI_uData_arShotSet{4}_SwitchOff_Pressure" : Real = PLC DB_MouldEditor_HMI.uData.arShotSet[4].SwitchOff_Pressure AT %DB10.DBD396, 1 s
   "DB_MouldEditor_HMI_uData_arShotSet{4}_RefComponent" : Int = PLC DB_MouldEditor_HMI.uData.arShotSet[4].RefComponent AT %DB10.DBW450, 1 s
   "DB_MouldEditor_HMI_uData_arShotSet{4}_2PoinMovement_Comp01" : Bool = PLC DB_MouldEditor_HMI.uData.arShotSet[4].2PoinMovement_Comp01 AT %DB10.DBX452.3, 1 s
   "DB_MouldEditor_HMI_uData_arShotSet{4}_2PoinMovement_Comp02" : Bool = PLC DB_MouldEditor_HMI.uData.arShotSet[4].2PoinMovement_Comp02 AT %DB10.DBX452.4, 1 s
   "DB_MouldEditor_HMI_uData_arShotSet{4}_2PoinMovement_Comp03" : Bool = PLC DB_MouldEditor_HMI.uData.arShotSet[4].2PoinMovement_Comp03 AT %DB10.DBX452.5, 1 s
   "DB_MouldEditor_HMI_uData_arShotSet{4}_2PoinMovement_Comp04" : Bool = PLC DB_MouldEditor_HMI.uData.arShotSet[4].2PoinMovement_Comp04 AT %DB10.DBX452.6, 1 s
   "DB_MouldEditor_HMI_uData_arShotSet{4}_2PoinMovement_Comp05" : Bool = PLC DB_MouldEditor_HMI.uData.arShotSet[4].2PoinMovement_Comp05 AT %DB10.DBX452.7, 1 s
   "DB_MouldEditor_HMI_uData_arShotSet{4}_2PoinMovement_Comp06" : Bool = PLC DB_MouldEditor_HMI.uData.arShotSet[4].2PoinMovement_Comp06 AT %DB10.DBX453.0, 1 s
   "DB_MouldEditor_HMI_uData_arShotSet{4}_Spare_1" : Bool = PLC DB_MouldEditor_HMI.uData.arShotSet[4].Spare_1 AT %DB10.DBX453.1, 1 s
   "DB_MouldEditor_HMI_uData_arShotSet{4}_Spare_2" : Bool = PLC DB_MouldEditor_HMI.uData.arShotSet[4].Spare_2 AT %DB10.DBX453.2, 1 s
   "DB_MouldEditor_HMI_uData_arShotSet{4}_Spare_3" : Bool = PLC DB_MouldEditor_HMI.uData.arShotSet[4].Spare_3 AT %DB10.DBX453.3, 1 s
   "DB_MouldEditor_HMI_uData_arShotSet{4}_Spare_4" : Bool = PLC DB_MouldEditor_HMI.uData.arShotSet[4].Spare_4 AT %DB10.DBX453.4, 1 s
   "DB_MouldEditor_HMI_uData_arShotSet{4}_Spare_5" : Bool = PLC DB_MouldEditor_HMI.uData.arShotSet[4].Spare_5 AT %DB10.DBX453.5, 1 s
   "DB_MouldEditor_HMI_uData_arShotSet{4}_Spare_6" : Bool = PLC DB_MouldEditor_HMI.uData.arShotSet[4].Spare_6 AT %DB10.DBX453.6, 1 s
   "DB_MouldEditor_HMI_uData_arShotSet{4}_Spare_7" : Bool = PLC DB_MouldEditor_HMI.uData.arShotSet[4].Spare_7 AT %DB10.DBX453.7, 1 s
   "DB_MouldEditor_HMI_uData_arShotSet{5}_CP_ThrottleGap" : Real = PLC DB_MouldEditor_HMI.uData.arShotSet[5].CP_ThrottleGap AT %DB10.DBD464, 1 s
   "DB_MouldEditor_HMI_uData_arShotSet{5}_SwitchOff_Pressure" : Real = PLC DB_MouldEditor_HMI.uData.arShotSet[5].SwitchOff_Pressure AT %DB10.DBD468, 1 s
   "DB_MouldEditor_HMI_uData_arShotSet{5}_RefComponent" : Int = PLC DB_MouldEditor_HMI.uData.arShotSet[5].RefComponent AT %DB10.DBW522, 1 s
   "DB_MouldEditor_HMI_uData_arShotSet{5}_2PoinMovement_Comp01" : Bool = PLC DB_MouldEditor_HMI.uData.arShotSet[5].2PoinMovement_Comp01 AT %DB10.DBX524.3, 1 s
   "DB_MouldEditor_HMI_uData_arShotSet{5}_2PoinMovement_Comp02" : Bool = PLC DB_MouldEditor_HMI.uData.arShotSet[5].2PoinMovement_Comp02 AT %DB10.DBX524.4, 1 s
   "DB_MouldEditor_HMI_uData_arShotSet{5}_2PoinMovement_Comp03" : Bool = PLC DB_MouldEditor_HMI.uData.arShotSet[5].2PoinMovement_Comp03 AT %DB10.DBX524.5, 1 s
   "DB_MouldEditor_HMI_uData_arShotSet{5}_2PoinMovement_Comp04" : Bool = PLC DB_MouldEditor_HMI.uData.arShotSet[5].2PoinMovement_Comp04 AT %DB10.DBX524.6, 1 s
   "DB_MouldEditor_HMI_uData_arShotSet{5}_2PoinMovement_Comp05" : Bool = PLC DB_MouldEditor_HMI.uData.arShotSet[5].2PoinMovement_Comp05 AT %DB10.DBX524.7, 1 s
   "DB_MouldEditor_HMI_uData_arShotSet{5}_2PoinMovement_Comp06" : Bool = PLC DB_MouldEditor_HMI.uData.arShotSet[5].2PoinMovement_Comp06 AT %DB10.DBX525.0, 1 s
   "DB_MouldEditor_HMI_uData_arShotSet{5}_Spare_1" : Bool = PLC DB_MouldEditor_HMI.uData.arShotSet[5].Spare_1 AT %DB10.DBX525.1, 1 s
   "DB_MouldEditor_HMI_uData_arShotSet{5}_Spare_2" : Bool = PLC DB_MouldEditor_HMI.uData.arShotSet[5].Spare_2 AT %DB10.DBX525.2, 1 s
   "DB_MouldEditor_HMI_uData_arShotSet{5}_Spare_3" : Bool = PLC DB_MouldEditor_HMI.uData.arShotSet[5].Spare_3 AT %DB10.DBX525.3, 1 s
   "DB_MouldEditor_HMI_uData_arShotSet{5}_Spare_4" : Bool = PLC DB_MouldEditor_HMI.uData.arShotSet[5].Spare_4 AT %DB10.DBX525.4, 1 s
   "DB_MouldEditor_HMI_uData_arShotSet{5}_Spare_5" : Bool = PLC DB_MouldEditor_HMI.uData.arShotSet[5].Spare_5 AT %DB10.DBX525.5, 1 s
   "DB_MouldEditor_HMI_uData_arShotSet{5}_Spare_6" : Bool = PLC DB_MouldEditor_HMI.uData.arShotSet[5].Spare_6 AT %DB10.DBX525.6, 1 s
   "DB_MouldEditor_HMI_uData_arShotSet{5}_Spare_7" : Bool = PLC DB_MouldEditor_HMI.uData.arShotSet[5].Spare_7 AT %DB10.DBX525.7, 1 s
   "DB_MouldEditor_HMI_uData_arShotSet{6}_CP_ThrottleGap" : Real = PLC DB_MouldEditor_HMI.uData.arShotSet[6].CP_ThrottleGap AT %DB10.DBD536, 1 s
   "DB_MouldEditor_HMI_uData_arShotSet{6}_SwitchOff_Pressure" : Real = PLC DB_MouldEditor_HMI.uData.arShotSet[6].SwitchOff_Pressure AT %DB10.DBD540, 1 s
   "DB_MouldEditor_HMI_uData_arShotSet{6}_RefComponent" : Int = PLC DB_MouldEditor_HMI.uData.arShotSet[6].RefComponent AT %DB10.DBW594, 1 s
   "DB_MouldEditor_HMI_uData_arShotSet{6}_2PoinMovement_Comp01" : Bool = PLC DB_MouldEditor_HMI.uData.arShotSet[6].2PoinMovement_Comp01 AT %DB10.DBX596.3, 1 s
   "DB_MouldEditor_HMI_uData_arShotSet{6}_2PoinMovement_Comp02" : Bool = PLC DB_MouldEditor_HMI.uData.arShotSet[6].2PoinMovement_Comp02 AT %DB10.DBX596.4, 1 s
   "DB_MouldEditor_HMI_uData_arShotSet{6}_2PoinMovement_Comp03" : Bool = PLC DB_MouldEditor_HMI.uData.arShotSet[6].2PoinMovement_Comp03 AT %DB10.DBX596.5, 1 s
   "DB_MouldEditor_HMI_uData_arShotSet{6}_2PoinMovement_Comp04" : Bool = PLC DB_MouldEditor_HMI.uData.arShotSet[6].2PoinMovement_Comp04 AT %DB10.DBX596.6, 1 s
   "DB_MouldEditor_HMI_uData_arShotSet{6}_2PoinMovement_Comp05" : Bool = PLC DB_MouldEditor_HMI.uData.arShotSet[6].2PoinMovement_Comp05 AT %DB10.DBX596.7, 1 s
   "DB_MouldEditor_HMI_uData_arShotSet{6}_2PoinMovement_Comp06" : Bool = PLC DB_MouldEditor_HMI.uData.arShotSet[6].2PoinMovement_Comp06 AT %DB10.DBX597.0, 1 s
   "DB_MouldEditor_HMI_uData_arShotSet{6}_Spare_1" : Bool = PLC DB_MouldEditor_HMI.uData.arShotSet[6].Spare_1 AT %DB10.DBX597.1, 1 s
   "DB_MouldEditor_HMI_uData_arShotSet{6}_Spare_2" : Bool = PLC DB_MouldEditor_HMI.uData.arShotSet[6].Spare_2 AT %DB10.DBX597.2, 1 s
   "DB_MouldEditor_HMI_uData_arShotSet{6}_Spare_3" : Bool = PLC DB_MouldEditor_HMI.uData.arShotSet[6].Spare_3 AT %DB10.DBX597.3, 1 s
   "DB_MouldEditor_HMI_uData_arShotSet{6}_Spare_4" : Bool = PLC DB_MouldEditor_HMI.uData.arShotSet[6].Spare_4 AT %DB10.DBX597.4, 1 s
   "DB_MouldEditor_HMI_uData_arShotSet{6}_Spare_5" : Bool = PLC DB_MouldEditor_HMI.uData.arShotSet[6].Spare_5 AT %DB10.DBX597.5, 1 s
   "DB_MouldEditor_HMI_uData_arShotSet{6}_Spare_6" : Bool = PLC DB_MouldEditor_HMI.uData.arShotSet[6].Spare_6 AT %DB10.DBX597.6, 1 s
   "DB_MouldEditor_HMI_uData_arShotSet{6}_Spare_7" : Bool = PLC DB_MouldEditor_HMI.uData.arShotSet[6].Spare_7 AT %DB10.DBX597.7, 1 s
   "DB_MouldEditor_HMI_uData_arShotSet{7}_CP_ThrottleGap" : Real = PLC DB_MouldEditor_HMI.uData.arShotSet[7].CP_ThrottleGap AT %DB10.DBD608, 1 s
   "DB_MouldEditor_HMI_uData_arShotSet{7}_SwitchOff_Pressure" : Real = PLC DB_MouldEditor_HMI.uData.arShotSet[7].SwitchOff_Pressure AT %DB10.DBD612, 1 s
   "DB_MouldEditor_HMI_uData_arShotSet{7}_RefComponent" : Int = PLC DB_MouldEditor_HMI.uData.arShotSet[7].RefComponent AT %DB10.DBW666, 1 s
   "DB_MouldEditor_HMI_uData_arShotSet{7}_2PoinMovement_Comp01" : Bool = PLC DB_MouldEditor_HMI.uData.arShotSet[7].2PoinMovement_Comp01 AT %DB10.DBX668.3, 1 s
   "DB_MouldEditor_HMI_uData_arShotSet{7}_2PoinMovement_Comp02" : Bool = PLC DB_MouldEditor_HMI.uData.arShotSet[7].2PoinMovement_Comp02 AT %DB10.DBX668.4, 1 s
   "DB_MouldEditor_HMI_uData_arShotSet{7}_2PoinMovement_Comp03" : Bool = PLC DB_MouldEditor_HMI.uData.arShotSet[7].2PoinMovement_Comp03 AT %DB10.DBX668.5, 1 s
   "DB_MouldEditor_HMI_uData_arShotSet{7}_2PoinMovement_Comp04" : Bool = PLC DB_MouldEditor_HMI.uData.arShotSet[7].2PoinMovement_Comp04 AT %DB10.DBX668.6, 1 s
   "DB_MouldEditor_HMI_uData_arShotSet{7}_2PoinMovement_Comp05" : Bool = PLC DB_MouldEditor_HMI.uData.arShotSet[7].2PoinMovement_Comp05 AT %DB10.DBX668.7, 1 s
   "DB_MouldEditor_HMI_uData_arShotSet{7}_2PoinMovement_Comp06" : Bool = PLC DB_MouldEditor_HMI.uData.arShotSet[7].2PoinMovement_Comp06 AT %DB10.DBX669.0, 1 s
   "DB_MouldEditor_HMI_uData_arShotSet{7}_Spare_1" : Bool = PLC DB_MouldEditor_HMI.uData.arShotSet[7].Spare_1 AT %DB10.DBX669.1, 1 s
   "DB_MouldEditor_HMI_uData_arShotSet{7}_Spare_2" : Bool = PLC DB_MouldEditor_HMI.uData.arShotSet[7].Spare_2 AT %DB10.DBX669.2, 1 s
   "DB_MouldEditor_HMI_uData_arShotSet{7}_Spare_3" : Bool = PLC DB_MouldEditor_HMI.uData.arShotSet[7].Spare_3 AT %DB10.DBX669.3, 1 s
   "DB_MouldEditor_HMI_uData_arShotSet{7}_Spare_4" : Bool = PLC DB_MouldEditor_HMI.uData.arShotSet[7].Spare_4 AT %DB10.DBX669.4, 1 s
   "DB_MouldEditor_HMI_uData_arShotSet{7}_Spare_5" : Bool = PLC DB_MouldEditor_HMI.uData.arShotSet[7].Spare_5 AT %DB10.DBX669.5, 1 s
   "DB_MouldEditor_HMI_uData_arShotSet{7}_Spare_6" : Bool = PLC DB_MouldEditor_HMI.uData.arShotSet[7].Spare_6 AT %DB10.DBX669.6, 1 s
   "DB_MouldEditor_HMI_uData_arShotSet{7}_Spare_7" : Bool = PLC DB_MouldEditor_HMI.uData.arShotSet[7].Spare_7 AT %DB10.DBX669.7, 1 s
   "DB_MouldEditor_HMI_uData_arShotSet{8}_CP_ThrottleGap" : Real = PLC DB_MouldEditor_HMI.uData.arShotSet[8].CP_ThrottleGap AT %DB10.DBD680, 1 s
   "DB_MouldEditor_HMI_uData_arShotSet{8}_SwitchOff_Pressure" : Real = PLC DB_MouldEditor_HMI.uData.arShotSet[8].SwitchOff_Pressure AT %DB10.DBD684, 1 s
   "DB_MouldEditor_HMI_uData_arShotSet{8}_RefComponent" : Int = PLC DB_MouldEditor_HMI.uData.arShotSet[8].RefComponent AT %DB10.DBW738, 1 s
   "DB_MouldEditor_HMI_uData_arShotSet{8}_2PoinMovement_Comp01" : Bool = PLC DB_MouldEditor_HMI.uData.arShotSet[8].2PoinMovement_Comp01 AT %DB10.DBX740.3, 1 s
   "DB_MouldEditor_HMI_uData_arShotSet{8}_2PoinMovement_Comp02" : Bool = PLC DB_MouldEditor_HMI.uData.arShotSet[8].2PoinMovement_Comp02 AT %DB10.DBX740.4, 1 s
   "DB_MouldEditor_HMI_uData_arShotSet{8}_2PoinMovement_Comp03" : Bool = PLC DB_MouldEditor_HMI.uData.arShotSet[8].2PoinMovement_Comp03 AT %DB10.DBX740.5, 1 s
   "DB_MouldEditor_HMI_uData_arShotSet{8}_2PoinMovement_Comp04" : Bool = PLC DB_MouldEditor_HMI.uData.arShotSet[8].2PoinMovement_Comp04 AT %DB10.DBX740.6, 1 s
   "DB_MouldEditor_HMI_uData_arShotSet{8}_2PoinMovement_Comp05" : Bool = PLC DB_MouldEditor_HMI.uData.arShotSet[8].2PoinMovement_Comp05 AT %DB10.DBX740.7, 1 s
   "DB_MouldEditor_HMI_uData_arShotSet{8}_2PoinMovement_Comp06" : Bool = PLC DB_MouldEditor_HMI.uData.arShotSet[8].2PoinMovement_Comp06 AT %DB10.DBX741.0, 1 s
   "DB_MouldEditor_HMI_uData_arShotSet{8}_Spare_1" : Bool = PLC DB_MouldEditor_HMI.uData.arShotSet[8].Spare_1 AT %DB10.DBX741.1, 1 s
   "DB_MouldEditor_HMI_uData_arShotSet{8}_Spare_2" : Bool = PLC DB_MouldEditor_HMI.uData.arShotSet[8].Spare_2 AT %DB10.DBX741.2, 1 s
   "DB_MouldEditor_HMI_uData_arShotSet{8}_Spare_3" : Bool = PLC DB_MouldEditor_HMI.uData.arShotSet[8].Spare_3 AT %DB10.DBX741.3, 1 s
   "DB_MouldEditor_HMI_uData_arShotSet{8}_Spare_4" : Bool = PLC DB_MouldEditor_HMI.uData.arShotSet[8].Spare_4 AT %DB10.DBX741.4, 1 s
   "DB_MouldEditor_HMI_uData_arShotSet{8}_Spare_5" : Bool = PLC DB_MouldEditor_HMI.uData.arShotSet[8].Spare_5 AT %DB10.DBX741.5, 1 s
   "DB_MouldEditor_HMI_uData_arShotSet{8}_Spare_6" : Bool = PLC DB_MouldEditor_HMI.uData.arShotSet[8].Spare_6 AT %DB10.DBX741.6, 1 s
   "DB_MouldEditor_HMI_uData_arShotSet{8}_Spare_7" : Bool = PLC DB_MouldEditor_HMI.uData.arShotSet[8].Spare_7 AT %DB10.DBX741.7, 1 s
   "DB_MouldEditor_HMI_uData_arShotSet{0}_Pressure{1}" : Real = PLC DB_MouldEditor_HMI.uData.arShotSet[0].Pressure[1] AT %DB10.DBD114, 1 s
   "DB_MouldEditor_HMI_uData_arShotSet{0}_Pressure{2}" : Real = PLC DB_MouldEditor_HMI.uData.arShotSet[0].Pressure[2] AT %DB10.DBD118, 1 s
   "DB_MouldEditor_HMI_uData_arShotSet{0}_Pressure{3}" : Real = PLC DB_MouldEditor_HMI.uData.arShotSet[0].Pressure[3] AT %DB10.DBD122, 1 s